HMI tags "DB_SDC_EMS_PAR_DRIVE"
   "_Byte_EMS[XXX].DRIVE_Delay_Pos" : Int, internal   // Absolute Position / absolute Positon
   "_Byte_EMS[XXX].DRIVE_DelaySpeedContr" : Int, internal   // Absolute Position / absolute Positon
   "_Byte_EMS[XXX].DRIVE_DIV_POS_FAST" : Int, internal   // Absolute Position / absolute Positon
   "_Byte_EMS[XXX].DRIVE_DIV_POS_SLOW" : Int, internal   // Absolute Position / absolute Positon
   "_Byte_EMS[XXX].DRIVE_FUNCT" : Int, internal   // Absolute Position / absolute Positon
   "_Byte_EMS[XXX].DRIVE_TOL_RESET_POS" : Int, internal   // Absolute Position / absolute Positon
   "_Byte_EMS[XXX].DRIVE_TOL_SET_POS" : Int, internal   // Absolute Position / absolute Positon
   "_Byte_EMS[XXX].DRIVE_TolSpeedContr" : Int, internal   // Absolute Position / absolute Positon
   "_Byte_EMS[XXX].DRIVE_V_DIV_FAST" : Int, internal   // Absolute Position / absolute Positon
   "_Byte_EMS[XXX].DRIVE_V_FACT_1" : Int, internal   // Absolute Position / absolute Positon
   "_Byte_EMS[XXX].DRIVE_V_FACT_2" : Int, internal   // Absolute Position / absolute Positon
   "_Byte_EMS[XXX].DRIVE_V_FACT_3" : Int, internal   // Absolute Position / absolute Positon
   "_Byte_EMS[XXX].DRIVE_V_FACT_4" : Int, internal   // Absolute Position / absolute Positon
   "_Byte_EMS[XXX].DRIVE_V_FACT_5" : Int, internal   // Absolute Position / absolute Positon
   "_Byte_EMS[XXX].DRIVE_V_Fixed_1" : Int, internal   // Absolute Position / absolute Positon
   "_Byte_EMS[XXX].DRIVE_V_Fixed_2" : Int, internal   // Absolute Position / absolute Positon
   "_Byte_EMS[XXX].DRIVE_V_Fixed_4_SLS_SPEED" : Int, internal   // Absolute Position / absolute Positon
   "_Byte_EMS[XXX].DRIVE_V_LIMIT_FACT" : Int, internal   // Absolute Position / absolute Positon
   "_Byte_EMS[XXX].DRIVE_V_max_Not_top" : Int, internal   // Absolute Position / absolute Positon
   "_Byte_EMS[XXX].DRIVE_V_max_top" : Int, internal   // Absolute Position / absolute Positon
   "_Byte_EMS[XXX].DRIVE_V_min" : Int, internal   // Absolute Position / absolute Positon
   "_Byte_EMS[XXX].DRIVE_V_Pos_2" : Int, internal   // Absolute Position / absolute Positon
   "_Byte_EMS[XXX].DRIVE_V_SETP_1" : Int, internal   // Absolute Position / absolute Positon
   "_Byte_EMS[XXX].DRIVE_V_SETP_2" : Int, internal   // Absolute Position / absolute Positon
   "_Byte_EMS[XXX].DRIVE_V_SETP_3" : Int, internal   // Absolute Position / absolute Positon
   "_Byte_EMS[XXX].DRIVE_V_SETP_4" : Int, internal   // Absolute Position / absolute Positon
   "_Byte_EMS[XXX].DRIVE_Window_Movement" : Int, internal   // Absolute Position / absolute Positon
   "_Byte_EMS[XXX].DRIVE_Window_Overrun" : Int, internal   // Absolute Position / absolute Positon
   "_Byte_EMS[XXX].DRIVE_Window_Pos" : Int, internal   // Absolute Position / absolute Positon
   "_Byte_EMS[XXX].DRIVE_Window_Pos_2" : Int, internal   // Absolute Position / absolute Positon
   "DB_SDC_EMS_PAR_HMI.HMI[XX].PAR.DRIVE.Delay_Pos" : Int AT %DB0.DBW0, 1 s
   "DB_SDC_EMS_PAR_HMI.HMI[XX].PAR.DRIVE.DelaySpeedContr" : S5Time AT %DB0.DBW0, 1 s
   "DB_SDC_EMS_PAR_HMI.HMI[XX].PAR.DRIVE.DIV_POS_FAST" : DInt AT %DB0.DBD0, 1 s
   "DB_SDC_EMS_PAR_HMI.HMI[XX].PAR.DRIVE.DIV_POS_SLOW" : DInt AT %DB0.DBD0, 1 s
   "DB_SDC_EMS_PAR_HMI.HMI[XX].PAR.DRIVE.TOL_RESET_POS" : Int AT %DB0.DBW0, 1 s
   "DB_SDC_EMS_PAR_HMI.HMI[XX].PAR.DRIVE.TOL_SET_POS" : Int AT %DB0.DBW0, 1 s
   "DB_SDC_EMS_PAR_HMI.HMI[XX].PAR.DRIVE.TolSpeedContr" : Int AT %DB0.DBW0, 1 s
   "DB_SDC_EMS_PAR_HMI.HMI[XX].PAR.DRIVE.V_DIV_FAST" : DInt AT %DB0.DBD0, 1 s
   "DB_SDC_EMS_PAR_HMI.HMI[XX].PAR.DRIVE.V_Fixed_1" : DInt AT %DB0.DBD0, 1 s
   "DB_SDC_EMS_PAR_HMI.HMI[XX].PAR.DRIVE.V_Fixed_2" : DInt AT %DB0.DBD0, 1 s
   "DB_SDC_EMS_PAR_HMI.HMI[XX].PAR.DRIVE.V_Fixed_4_SLS_SPEED" : DInt AT %DB0.DBD0, 1 s
   "DB_SDC_EMS_PAR_HMI.HMI[XX].PAR.DRIVE.V_max_Not_top" : DInt AT %DB0.DBD0, 1 s
   "DB_SDC_EMS_PAR_HMI.HMI[XX].PAR.DRIVE.V_max_top" : DInt AT %DB0.DBD0, 1 s
   "DB_SDC_EMS_PAR_HMI.HMI[XX].PAR.DRIVE.V_min" : DInt AT %DB0.DBD0, 1 s
   "DB_SDC_EMS_PAR_HMI.HMI[XX].PAR.DRIVE.V_Pos_2" : DInt AT %DB0.DBD0, 1 s
   "DB_SDC_EMS_PAR_HMI.HMI[XX].PAR.DRIVE.Window_Movement" : Int AT %DB0.DBW0, 1 s
   "DB_SDC_EMS_PAR_HMI.HMI[XX].PAR.DRIVE.Window_Overrun" : Int AT %DB0.DBW0, 1 s
   "DB_SDC_EMS_PAR_HMI.HMI[XX].PAR.DRIVE.Window_Pos" : Int AT %DB0.DBW0, 1 s
   "DB_SDC_EMS_PAR_HMI.HMI[XX].PAR.DRIVE.Window_Pos_2" : Int AT %DB0.DBW0, 1 s
   "DB_SDC_EMS_PAR_HMI.HMI[XX].PAR.DRIVE.Funct" : Word AT %DB0.DBW0, 1 s
   "DB_SDC_EMS_PAR_HMI.HMI[XX].PAR.DRIVE.V_FACT_1" : Real AT %DB0.DBD0, 1 s
   "DB_SDC_EMS_PAR_HMI.HMI[XX].PAR.DRIVE.V_FACT_2" : Real AT %DB0.DBD0, 1 s
   "DB_SDC_EMS_PAR_HMI.HMI[XX].PAR.DRIVE.V_FACT_3" : Real AT %DB0.DBD0, 1 s
   "DB_SDC_EMS_PAR_HMI.HMI[XX].PAR.DRIVE.V_FACT_4" : Real AT %DB0.DBD0, 1 s
   "DB_SDC_EMS_PAR_HMI.HMI[XX].PAR.DRIVE.V_FACT_5" : Real AT %DB0.DBD0, 1 s
   "DB_SDC_EMS_PAR_HMI.HMI[XX].PAR.DRIVE.V_LIMIT_FACT" : Real AT %DB0.DBD0, 1 s
   "DB_SDC_EMS_PAR_HMI.HMI[XX].PAR.DRIVE.V_SETP_1" : DInt AT %DB0.DBD0, 1 s
   "DB_SDC_EMS_PAR_HMI.HMI[XX].PAR.DRIVE.V_SETP_2" : DInt AT %DB0.DBD0, 1 s
   "DB_SDC_EMS_PAR_HMI.HMI[XX].PAR.DRIVE.V_SETP_3" : DInt AT %DB0.DBD0, 1 s
   "DB_SDC_EMS_PAR_HMI.HMI[XX].PAR.DRIVE.V_SETP_4" : DInt AT %DB0.DBD0, 1 s
   "_Byte_EMS[XXX].DRIVE_Delay_Pos(1)" : Int, internal

HMI tags "DB_SDC_EMS_PAR_HOIST"
   "_Byte_EMS[XXX].HOIST_V_min" : Int, internal   // Absolute Position / absolute Positon
   "DB_SDC_EMS_PAR_HMI.HMI[XX].PAR.HOIST.V_min" : Int AT %DB0.DBW0, 1 s
   "_Byte_EMS[XXX].HOIST_V_max" : Int, internal   // Absolute Position / absolute Positon
   "DB_SDC_EMS_PAR_HMI.HMI[XX].PAR.HOIST.V_max" : Int AT %DB0.DBW0, 1 s
   "_Byte_EMS[XXX].HOIST_V_MaxOccLift" : Int, internal   // Absolute Position / absolute Positon
   "DB_SDC_EMS_PAR_HMI.HMI[XX].PAR.HOIST.V_MaxOccLift" : Int AT %DB0.DBW0, 1 s
   "_Byte_EMS[XXX].HOIST_V_Pos_1" : Int, internal   // Absolute Position / absolute Positon
   "DB_SDC_EMS_PAR_HMI.HMI[XX].PAR.HOIST.V_Pos_1" : Int AT %DB0.DBW0, 1 s
   "_Byte_EMS[XXX].HOIST_V_Pos_2" : Int, internal   // Absolute Position / absolute Positon
   "DB_SDC_EMS_PAR_HMI.HMI[XX].PAR.HOIST.V_Pos_2" : Int AT %DB0.DBW0, 1 s
   "_Byte_EMS[XXX].HOIST_V_Fixed_1" : Int, internal   // Absolute Position / absolute Positon
   "DB_SDC_EMS_PAR_HMI.HMI[XX].PAR.HOIST.V_Fixed_1" : Int AT %DB0.DBW0, 1 s
   "_Byte_EMS[XXX].HOIST_V_Fixed_2" : Int, internal   // Absolute Position / absolute Positon
   "DB_SDC_EMS_PAR_HMI.HMI[XX].PAR.HOIST.V_Fixed_2" : Int AT %DB0.DBW0, 1 s
   "_Byte_EMS[XXX].HOIST_V_Fixed_4" : Int, internal   // Absolute Position / absolute Positon
   "DB_SDC_EMS_PAR_HMI.HMI[XX].PAR.HOIST.V_Fixed_4" : Int AT %DB0.DBW0, 1 s
   "_Byte_EMS[XXX].HOIST_V_Fixed_6" : Int, internal   // Absolute Position / absolute Positon
   "DB_SDC_EMS_PAR_HMI.HMI[XX].PAR.HOIST.V_Fixed_6" : Int AT %DB0.DBW0, 1 s
   "_Byte_EMS[XXX].HOIST_V_FACT_Hz_UP" : Int, internal   // Absolute Position / absolute Positon
   "DB_SDC_EMS_PAR_HMI.HMI[XX].PAR.HOIST.V_FACT_Hz_UP" : Real AT %DB0.DBD0, 1 s
   "_Byte_EMS[XXX].HOIST_V_FACT_Hz_DOWN" : Int, internal   // Absolute Position / absolute Positon
   "DB_SDC_EMS_PAR_HMI.HMI[XX].PAR.HOIST.V_FACT_Hz_DOWN" : Real AT %DB0.DBD0, 1 s
   "DB_SDC_EMS_PAR_HMI.HMI[XX].PAR.HOIST.H_Window_POS_V1" : Int AT %DB0.DBW0, 1 s
   "_Byte_EMS[XXX].HOIST_H_Window_POS_V1" : Int, internal   // Absolute Position / absolute Positon
   "DB_SDC_EMS_PAR_HMI.HMI[XX].PAR.HOIST.H_Window_POS_V2" : Int AT %DB0.DBW0, 1 s
   "_Byte_EMS[XXX].HOIST_H_Window_POS_V2" : Int, internal   // Absolute Position / absolute Positon
   "DB_SDC_EMS_PAR_HMI.HMI[XX].PAR.HOIST.H_TOL_SET_POS" : Int AT %DB0.DBW0, 1 s
   "_Byte_EMS[XXX].HOIST_H_TOL_SET_POS" : Int, internal   // Absolute Position / absolute Positon
   "DB_SDC_EMS_PAR_HMI.HMI[XX].PAR.HOIST.H_TOL_RESET_POS" : Int AT %DB0.DBW0, 1 s
   "_Byte_EMS[XXX].HOIST_H_TOL_RESET_POS" : Int, internal   // Absolute Position / absolute Positon
   "DB_SDC_EMS_PAR_HMI.HMI[XX].PAR.HOIST.H_MIN" : Int AT %DB0.DBW0, 1 s
   "_Byte_EMS[XXX].HOIST_H_MIN" : Int, internal   // Absolute Position / absolute Positon
   "DB_SDC_EMS_PAR_HMI.HMI[XX].PAR.HOIST.H_MIN_without_bypass" : Int AT %DB0.DBW0, 1 s
   "_Byte_EMS[XXX].HOIST_H_MIN_without_bypass" : Int, internal   // Absolute Position / absolute Positon
   "DB_SDC_EMS_PAR_HMI.HMI[XX].PAR.HOIST.H_REF_OFFSET" : Int AT %DB0.DBW0, 1 s
   "_Byte_EMS[XXX].HOIST_H_REF_OFFSET" : Int, internal   // Absolute Position / absolute Positon
   "DB_SDC_EMS_PAR_HMI.HMI[XX].PAR.HOIST.H_REF" : Int AT %DB0.DBW0, 1 s
   "_Byte_EMS[XXX].HOIST_H_REF" : Int, internal   // Absolute Position / absolute Positon
   "DB_SDC_EMS_PAR_HMI.HMI[XX].PAR.HOIST.H_FACT_ENC1" : Real AT %DB0.DBD0, 1 s
   "_Byte_EMS[XXX].HOIST_H_FACT_ENC1" : Int, internal   // Absolute Position / absolute Positon
   "DB_SDC_EMS_PAR_HMI.HMI[XX].PAR.HOIST.H_FACT_ENC2" : Real AT %DB0.DBD0, 1 s
   "_Byte_EMS[XXX].HOIST_H_FACT_ENC2" : Int, internal   // Absolute Position / absolute Positon
   "DB_SDC_EMS_PAR_HMI.HMI[XX].PAR.HOIST.H_FACT_SPEED" : Real AT %DB0.DBD0, 1 s
   "_Byte_EMS[XXX].HOIST_H_FACT_SPEED" : Int, internal   // Absolute Position / absolute Positon
   "DB_SDC_EMS_PAR_HMI.HMI[XX].PAR.HOIST.H_ENC_MAX_DIFF" : Int AT %DB0.DBW0, 1 s
   "_Byte_EMS[XXX].HOIST_H_ENC_MAX_DIFF" : Int, internal   // Absolute Position / absolute Positon
   "DB_SDC_EMS_PAR_HMI.HMI[XX].PAR.HOIST.H_Slow" : Int AT %DB0.DBW0, 1 s
   "_Byte_EMS[XXX].HOIST_H_Slow" : Int, internal   // Absolute Position / absolute Positon
   "DB_SDC_EMS_PAR_HMI.HMI[XX].PAR.HOIST.H_tIN_POS" : Int AT %DB0.DBW0, 1 s
   "_Byte_EMS[XXX].HOIST_H_tIN_POS" : Int, internal   // Absolute Position / absolute Positon
   "DB_SDC_EMS_PAR_HMI.HMI[XX].PAR.HOIST.H_REF_HMI" : Int AT %DB0.DBW0, 1 s
   "_Byte_EMS[XXX].HOIST_H_REF_HMI" : Int, internal   // Absolute Position / absolute Positon
   "_Byte_EMS[XXX].HOIST_V_Fixed_3" : Int, internal
   "DB_SDC_EMS_PAR_HMI.HMI[XX].PAR.HOIST.V_Fixed_3" : Int AT %DB0.DBW0, 1 s

HMI tags "VAT_SYSTEM_ALLG"
   "_intern_BILD_Nr" : Int, internal
   "_intern_1_bool" : Bool, internal
   "_intern_0_bool" : Bool, internal
   "_intern_1" : Int, internal
   "_intern_2" : Int, internal
   "_intern_3" : Int, internal
   "_intern_4" : Int, internal
   "_intern_5" : Int, internal
   "_intern_6" : Int, internal
   "_intern_7" : Int, internal
   "_intern_8" : Int, internal
   "_intern_9" : Int, internal
   "_intern_10" : Int, internal
   "_intern_11" : Int, internal
   "_intern_12" : Int, internal
   "_intern_13" : Int, internal
   "_intern_14" : Int, internal
   "_intern_15" : Int, internal
   "_intern_16" : Int, internal
   "_intern_17" : Int, internal
   "_intern_18" : Int, internal
   "_intern_19" : Int, internal
   "_intern_20" : Int, internal
   "_intern_21" : Int, internal
   "_intern_22" : Int, internal
   "_intern_23" : Int, internal
   "_intern_24" : Int, internal
   "_intern_25" : Int, internal
   "_intern_26" : Int, internal
   "_intern_27" : Int, internal
   "_intern_28" : Int, internal
   "_intern_29" : Int, internal
   "_intern_30" : Int, internal
   "_intern_31" : Int, internal
   "_intern_32" : Int, internal
   "_intern_33" : Int, internal
   "_intern_34" : Int, internal
   "_intern_35" : Int, internal
   "_intern_36" : Int, internal
   "_intern_37" : Int, internal
   "_intern_38" : Int, internal
   "_intern_39" : Int, internal
   "_intern_40" : Int, internal
   "_intern_41" : Int, internal
   "_intern_42" : Int, internal
   "_intern_43" : Int, internal
   "_intern_44" : Int, internal
   "_intern_45" : Int, internal
   "_intern_46" : Int, internal
   "_intern_47" : Int, internal
   "_intern_48" : Int, internal
   "_intern_49" : Int, internal
   "_intern_50" : Int, internal
   "_intern_51" : Int, internal
   "_intern_52" : Int, internal
   "_intern_53" : Int, internal
   "_intern_54" : Int, internal
   "_intern_55" : Int, internal
   "_intern_56" : Int, internal
   "_intern_57" : Int, internal
   "_intern_58" : Int, internal
   "_intern_59" : Int, internal
   "_intern_60" : Int, internal
   "_intern_61" : Int, internal
   "_intern_62" : Int, internal
   "_intern_63" : Int, internal
   "_intern_64" : Int, internal
   "_intern_65" : Int, internal
   "_intern_66" : Int, internal
   "_intern_67" : Int, internal
   "_intern_68" : Int, internal
   "_intern_69" : Int, internal
   "_intern_70" : Int, internal
   "_intern_71" : Int, internal
   "_intern_72" : Int, internal
   "_intern_73" : Int, internal
   "_intern_74" : Int, internal
   "_intern_75" : Int, internal
   "_intern_76" : Int, internal
   "_intern_77" : Int, internal
   "_intern_78" : Int, internal
   "_intern_79" : Int, internal
   "_intern_80" : Int, internal
   "_intern_81" : Int, internal
   "_intern_82" : Int, internal
   "_intern_83" : Int, internal
   "_intern_84" : Int, internal
   "_intern_85" : Int, internal
   "_intern_86" : Int, internal
   "_intern_87" : Int, internal
   "_intern_88" : Int, internal
   "_intern_89" : Int, internal
   "_intern_90" : Int, internal
   "_intern_91" : Int, internal
   "_intern_92" : Int, internal
   "_intern_93" : Int, internal
   "_intern_94" : Int, internal
   "_intern_95" : Int, internal
   "_intern_96" : Int, internal
   "_intern_97" : Int, internal
   "_intern_98" : Int, internal
   "_intern_99" : Int, internal
   "_intern_100" : Int, internal
   "_intern_101" : Int, internal
   "_intern_102" : Int, internal
   "_intern_103" : Int, internal
   "_intern_104" : Int, internal
   "_intern_105" : Int, internal
   "_intern_106" : Int, internal
   "_intern_107" : Int, internal
   "_intern_108" : Int, internal
   "_intern_109" : Int, internal
   "_intern_110" : Int, internal
   "_intern_111" : Int, internal
   "_intern_112" : Int, internal
   "_intern_113" : Int, internal
   "_intern_114" : Int, internal
   "_intern_115" : Int, internal
   "_intern_116" : Int, internal
   "_intern_117" : Int, internal
   "_intern_118" : Int, internal
   "_intern_119" : Int, internal
   "_intern_120" : Int, internal
   "_intern_121" : Int, internal
   "_intern_122" : Int, internal
   "_intern_123" : Int, internal
   "_intern_124" : Int, internal
   "_intern_125" : Int, internal
   "_intern_126" : Int, internal
   "_intern_127" : Int, internal
   "_intern_128" : Int, internal
   "_intern_129" : Int, internal
   "_intern_130" : Int, internal
   "_intern_131" : Int, internal
   "_intern_132" : Int, internal
   "_intern_133" : Int, internal
   "_intern_134" : Int, internal
   "_intern_135" : Int, internal
   "_intern_136" : Int, internal
   "_intern_137" : Int, internal
   "_intern_138" : Int, internal
   "_intern_139" : Int, internal
   "_intern_140" : Int, internal
   "_intern_141" : Int, internal
   "_intern_142" : Int, internal
   "_intern_143" : Int, internal
   "_intern_144" : Int, internal
   "_intern_145" : Int, internal
   "_intern_146" : Int, internal
   "_intern_147" : Int, internal
   "_intern_148" : Int, internal
   "_intern_149" : Int, internal
   "_intern_150" : Int, internal
   "_intern_151" : Int, internal
   "_intern_152" : Int, internal
   "_intern_153" : Int, internal
   "_intern_154" : Int, internal
   "_intern_155" : Int, internal
   "_intern_156" : Int, internal
   "_intern_157" : Int, internal
   "_intern_158" : Int, internal
   "_intern_159" : Int, internal
   "_intern_160" : Int, internal
   "_intern_161" : Int, internal
   "_intern_162" : Int, internal
   "_intern_163" : Int, internal
   "_intern_164" : Int, internal
   "_intern_165" : Int, internal
   "_intern_166" : Int, internal
   "_intern_167" : Int, internal
   "_intern_168" : Int, internal
   "_intern_169" : Int, internal
   "_intern_170" : Int, internal
   "_intern_171" : Int, internal
   "_intern_172" : Int, internal
   "_intern_173" : Int, internal
   "_intern_174" : Int, internal
   "_intern_175" : Int, internal
   "_intern_176" : Int, internal
   "_intern_177" : Int, internal
   "_intern_178" : Int, internal
   "_intern_179" : Int, internal
   "_intern_180" : Int, internal
   "_intern_181" : Int, internal
   "_intern_182" : Int, internal
   "_intern_183" : Int, internal
   "_intern_184" : Int, internal
   "_intern_185" : Int, internal
   "_intern_186" : Int, internal
   "_intern_187" : Int, internal
   "_intern_188" : Int, internal
   "_intern_189" : Int, internal
   "_intern_190" : Int, internal
   "_intern_191" : Int, internal
   "_intern_192" : Int, internal
   "_intern_193" : Int, internal
   "_intern_194" : Int, internal
   "_intern_195" : Int, internal
   "_intern_196" : Int, internal
   "_intern_197" : Int, internal
   "_intern_198" : Int, internal
   "_intern_199" : Int, internal
   "_intern_200" : Int, internal

HMI tags "VAT_PN_PB"
   "PN_PB\PTMUX_P_TLN17_32" : UInt, internal
   "PN_PB\PTMUX_P_TLN1_16" : UInt, internal
   "PN_PB\PTMUX_P_TLN129_144" : UInt, internal
   "PN_PB\DB_PN" : UInt, internal
   "PN_PB\PTMUX_P_TLN177_192" : UInt, internal
   "PN_PB\PTMUX_F_TLN241_256" : UInt, internal
   "PN_PB\IO_Sys_ID" : Int, internal
   "PN_PB\PTMUX_P_TLN225_240" : UInt, internal
   "PN_PB\PTMUX_P_TLN241_256" : UInt, internal
   "PN_PB\PTMUX_P_TLN193_208" : UInt, internal
   "PN_PB\PTMUX_F_TLN1_16" : UInt, internal
   "PN_PB\PTMUX_P_TLN209_224" : UInt, internal
   "PN_PB\PTMUX_F_TLN49_64" : UInt, internal
   "PN_PB\PTMUX_P_TLN113_128" : UInt, internal
   "PN_PB\PTMUX_F_TLN177_192" : UInt, internal
   "PN_PB\PTMUX_P_TLN49_64" : UInt, internal
   "PN_PB\PTMUX_F_TLN97_112" : UInt, internal
   "PN_PB\DB_PB" : UInt, internal
   "PN_PB\PTMUX_F_TLN81_96" : UInt, internal
   "PN_PB\PTMUX_F_TLN145_160" : UInt, internal
   "PN_PB\Diag_Art" : Int, internal
   "PN_PB\PTMUX_F_TLN113_128" : UInt, internal
   "PN_PB\PTMUX_P_TLN97_112" : UInt, internal
   "PN_PB\Teiln_Nr_Anz." : Int, internal
   "PN_PB\PTMUX_P_TLN33_48" : UInt, internal
   "PN_PB\PTMUX_F_TLN161_176" : UInt, internal
   "PN_PB\PTMUX_F_TLN193_208" : UInt, internal
   "PN_PB\PTMUX_P_TLN81_96" : UInt, internal
   "PN_PB\PTMUX_P_TLN65_80" : UInt, internal
   "PN_PB\PTMUX_F_TLN225_240" : UInt, internal
   "PN_PB\PTMUX_F_TLN17_32" : UInt, internal
   "PN_PB\PTMUX_F_TLN65_80" : UInt, internal
   "PN_PB\PTMUX_F_TLN209_224" : UInt, internal
   "PN_PB\PTMUX_F_TLN33_48" : UInt, internal
   "PN_PB\PTMUX_P_TLN145_160" : UInt, internal
   "PN_PB\PTMUX_P_TLN161_176" : UInt, internal
   "PN_PB\Teiln_Nr_Bez" : WString[20], internal
   "PN_PB\Teiln_Nr_Typ" : WString[12], internal
   "PN_PB\Teiln_Nr_Ort" : WString[12], internal
   "PN_PB\PTMUX_F_TLN129_144" : UInt, internal

HMI tags "VAT_SYSTEM_PN"
   "PN_PB\PN\TLN_P_161_176" : Word AT %DB0.DBW230, 100 ms
   "PN_PB\PN\TLN_F_241_256" : Word AT %DB0.DBW368, 100 ms
   "PN_PB\PN\TLN_P_33_48" : Word AT %DB0.DBW214, 100 ms
   "PN_PB\PN\TLN_F_49_64" : Word AT %DB0.DBW344, 100 ms
   "PN_PB\PN\TLN_F_81_96" : Word AT %DB0.DBW348, 100 ms
   "PN_PB\PN\TLN_P_225_240" : Word AT %DB0.DBW238, 100 ms
   "PN_PB\PN\TLN_P_177_192" : Word AT %DB0.DBW232, 100 ms
   "PN_PB\PN\TLN_F_17_32" : Word AT %DB0.DBW340, 100 ms
   "PN_PB\PN\TLN_F_225_240" : Word AT %DB0.DBW366, 100 ms
   "PN_PB\PN\TLN_F_33_48" : Word AT %DB0.DBW342, 100 ms
   "PN_PB\PN\TLN_P_97_112" : Word AT %DB0.DBW222, 100 ms
   "PN_PB\PN\TLN_P_129_144" : Word AT %DB0.DBW226, 100 ms
   "PN_PB\PN\Diag_Slave_Nr" : Int, internal
   "PN_PB\PN\TLN_F_113_128" : Word AT %DB0.DBW352, 100 ms
   "PN_PB\PN\TLN_F_97_112" : Word AT %DB0.DBW350, 100 ms
   "PN_PB\PN\TLN_P_145_160" : Word AT %DB0.DBW228, 100 ms
   "PN_PB\PN\TLN_F_145_160" : Word AT %DB0.DBW356, 100 ms
   "PN_PB\PN\TLN_P_113_128" : Word AT %DB0.DBW224, 100 ms
   "PN_PB\PN\IOSys_ID" : Int AT %DB0.DBW2, 200 ms
   "PN_PB\PN\TLN_F_129_144" : Word AT %DB0.DBW354, 100 ms
   "PN_PB\PN\TLN_F_161_176" : Word AT %DB0.DBW358, 100 ms
   "PN_PB\PN\TLN_F_1_16" : Word AT %DB0.DBW338, 100 ms
   "PN_PB\PN\TLN_P_1_16" : Word AT %DB0.DBW210, 100 ms
   "PN_PB\PN\TLN_P_65_80" : Word AT %DB0.DBW218, 100 ms
   "PN_PB\PN\TLN_F_209_224" : Word AT %DB0.DBW364, 100 ms
   "PN_PB\PN\TLN_F_65_80" : Word AT %DB0.DBW346, 100 ms
   "PN_PB\PN\TLN_P_193_208" : Word AT %DB0.DBW234, 100 ms
   "PN_PB\PN\TLN_P_81_96" : Word AT %DB0.DBW220, 100 ms
   "PN_PB\PN\TLN_P_209_224" : Word AT %DB0.DBW236, 100 ms
   "PN_PB\PN\TLN_P_17_32" : Word AT %DB0.DBW212, 100 ms
   "PN_PB\PN\TLN_P_49_64" : Word AT %DB0.DBW216, 100 ms
   "PN_PB\PN\TLN_P_241_256" : Word AT %DB0.DBW240, 100 ms
   "PN_PB\PN\TLN_F_193_208" : Word AT %DB0.DBW362, 100 ms
   "PN_PB\PN\TLN_F_177_192" : Word AT %DB0.DBW360, 100 ms
   "PN_PB\PN\Teiln_Nr" : Int AT %DB0.DBW4, 1 s
      on ChangeValue: "SDC_PN"()

HMI tags "VAT_SYSTEM_PB"
   "PN_PB\PB\TLN_F_65_80" : Word AT %DB0.DBW234, 100 ms
   "PN_PB\PB\TLN_F_113_128" : Word AT %DB0.DBW240, 100 ms
   "PN_PB\PB\IOSys_ID" : Int AT %DB0.DBW2, 200 ms
   "PN_PB\PB\TLN_P_81_96" : Word AT %DB0.DBW220, 100 ms
   "PN_PB\PB\TLN_F_81_96" : Word AT %DB0.DBW236, 100 ms
   "PN_PB\PB\TLN_F_49_64" : Word AT %DB0.DBW232, 100 ms
   "PN_PB\PB\TLN_P_113_128" : Word AT %DB0.DBW224, 100 ms
   "PN_PB\PB\TLN_F_33_48" : Word AT %DB0.DBW230, 100 ms
   "PN_PB\PB\TLN_P_65_80" : Word AT %DB0.DBW218, 100 ms
   "PN_PB\PB\TLN_P_49_64" : Word AT %DB0.DBW216, 100 ms
   "PN_PB\PB\TLN_F_1_16" : Word AT %DB0.DBW226, 100 ms
   "PN_PB\PB\TLN_P_17_32" : Word AT %DB0.DBW212, 100 ms
   "PN_PB\PB\TLN_P_33_48" : Word AT %DB0.DBW214, 100 ms
   "PN_PB\PB\TLN_P_1_16" : Word AT %DB0.DBW210, 100 ms
   "PN_PB\PB\TLN_F_17_32" : Word AT %DB0.DBW228, 100 ms
   "PN_PB\PB\TLN_F_97_112" : Word AT %DB0.DBW238, 100 ms
   "PN_PB\PB\TLN_P_97_112" : Word AT %DB0.DBW222, 100 ms
   "PN_PB\PB\Teiln_Nr" : Int AT %DB0.DBW4, 200 ms

HMI tags "VAT_SYSTEM_PARAMETER"
   "_intern_Pult_Nr" : Int, internal   // !!! VOR DEM LADEN EINSTELLEN !!!

HMI tags "UserDiag_TagTable"
   "UserDiag_HmiData_actIOSystem" : Int = PLC UserDiag_HmiData.actIOSystem, 1 s
   "UserDiag_HmiData_actDeviceOfScreen" : Int = PLC UserDiag_HmiData.actDeviceOfScreen, 1 s
   "UserDiag_HmiData_ioSlotDiagnosticsLoaded" : Bool = PLC UserDiag_HmiData.ioSlotDiagnosticsLoaded, 1 s
   "UserDiag_HmiData_actScreenDevices" : Int = PLC UserDiag_HmiData.actScreenDevices, 100 ms
   "UserDiag_HmiData_maxScreensDevices" : Int = PLC UserDiag_HmiData.maxScreensDevices, 1 s
   "UserDiag_HmiData_ackWaitTime" : Int = PLC UserDiag_HmiData.ackWaitTime, 1 s
   "UserDiag_HmiData_ackStates" : Bool = PLC UserDiag_HmiData.ackStates, 1 s
   "UserDiag_HmiData_actIOSystemData" : UserDiag_typeActIOSystem = PLC UserDiag_HmiData.actIOSystemData, 1 s
   "UserDiag_HmiData_actDeviceNumber" : UInt = PLC UserDiag_HmiData.actDeviceNumber, 1 s
   "UserDiag_HmiData_actDeviceName" : String[50] = PLC UserDiag_HmiData.actDeviceName, 1 s
   "UserDiag_HmiData_actIPAddress.ADDR" : Array [0..3] of Byte = PLC UserDiag_HmiData.actIPAddress.ADDR, 1 s
   "UserDiag_HmiData_ioSystemError" : Array [0..1] of Bool = PLC UserDiag_HmiData.ioSystemError AT %DB1.DBX0.0, 500 ms
   "UserDiag_HmiData_filterErrorDevices" : Bool = PLC UserDiag_HmiData.filterErrorDevices AT %DB1.DBX0.0, 500 ms
   "UserDiag_HmiData_errorAtLowerScreen" : Bool = PLC UserDiag_HmiData.errorAtLowerScreen, 500 ms
   "UserDiag_HmiData_errorAtUpperScreen" : Bool = PLC UserDiag_HmiData.errorAtUpperScreen AT %DB1.DBW0, 500 ms
   "ioSystem1" : Int AT %DB1.DBW0
   "ioSystem2" : Int AT %DB1.DBW0
   "ioSystem3" : Int AT %DB1.DBW0
   "DB_SDC_FAULTS" : Word = PLC DB101_DB_SDC_FAULTS.SDC_Fault AT %DB101.DBW0, 1 s

HMI tags "DB_SDC_FAULTS"
   "DB101_DB_SDC_FAULTS_SDC_Fault" : Word = PLC DB101_DB_SDC_FAULTS.SDC_Fault AT %DB101.DBW0, 1 s
   "DB101_DB_SDC_FAULTS_Carrier_Fault[15]" : Word = PLC DB101_DB_SDC_FAULTS.Carrier_Fault[15] AT %DB101.DBW30, 1 s
   "DB101_DB_SDC_FAULTS_Carrier_Fault[27]" : Word = PLC DB101_DB_SDC_FAULTS.Carrier_Fault[27] AT %DB101.DBW54, 1 s
   "DB101_DB_SDC_FAULTS_Carrier_Fault[31]" : Word = PLC DB101_DB_SDC_FAULTS.Carrier_Fault[31] AT %DB101.DBW62, 1 s
   "DB101_DB_SDC_FAULTS_Carrier_Fault[40]" : Word = PLC DB101_DB_SDC_FAULTS.Carrier_Fault[40] AT %DB101.DBW80, 1 s

HMI tags "DB_HMI_FAULTS"
   "DB302_HMI_Faults_SDC_Faults_0" : Int = PLC DB302_HMI_Faults.SDC_Faults_0, 1 s
   "DB302_HMI_Faults_SDC_Faults_1" : Int = PLC DB302_HMI_Faults.SDC_Faults_1, 1 s
   "DB302_HMI_Faults_SDC_Faults_2" : Int = PLC DB302_HMI_Faults.SDC_Faults_2, 1 s
   "DB302_HMI_Faults_SDC_Faults_3" : Int = PLC DB302_HMI_Faults.SDC_Faults_3, 1 s

HMI tags "EMS"
   "EMS" : UDT_System = PLC EMS AT %DB1.DBW0, 1 s

HMI tags "DeviceStates_Condition"
   "DB16_EMS_Status_EMS_DeviceStates.DeviceStates_Condition_HMI[2]" : Int = PLC DB16_EMS_Status.EMS_DeviceStates.DeviceStates_Condition_HMI[2], 1 s
   "DB16_EMS_Status_EMS_DeviceStates.DeviceStates_Condition_HMI[3]" : Int = PLC DB16_EMS_Status.EMS_DeviceStates.DeviceStates_Condition_HMI[3], 1 s
   "DB16_EMS_Status_EMS_DeviceStates.DeviceStates_Condition_HMI[4]" : Int = PLC DB16_EMS_Status.EMS_DeviceStates.DeviceStates_Condition_HMI[4], 1 s
   "DB16_EMS_Status_EMS_DeviceStates.DeviceStates_Condition_HMI[5]" : Int = PLC DB16_EMS_Status.EMS_DeviceStates.DeviceStates_Condition_HMI[5], 1 s
   "DB16_EMS_Status_EMS_DeviceStates.DeviceStates_Condition_HMI[6]" : Int = PLC DB16_EMS_Status.EMS_DeviceStates.DeviceStates_Condition_HMI[6], 1 s
   "DB16_EMS_Status_EMS_DeviceStates.DeviceStates_Condition_HMI[7]" : Int = PLC DB16_EMS_Status.EMS_DeviceStates.DeviceStates_Condition_HMI[7], 1 s
   "DB16_EMS_Status_EMS_DeviceStates.DeviceStates_Condition_HMI[8]" : Int = PLC DB16_EMS_Status.EMS_DeviceStates.DeviceStates_Condition_HMI[8], 1 s
   "DB16_EMS_Status_EMS_DeviceStates.DeviceStates_Condition_HMI[9]" : Int = PLC DB16_EMS_Status.EMS_DeviceStates.DeviceStates_Condition_HMI[9], 1 s
   "DB16_EMS_Status_EMS_DeviceStates.DeviceStates_Condition_HMI[10]" : Int = PLC DB16_EMS_Status.EMS_DeviceStates.DeviceStates_Condition_HMI[10], 1 s
   "DB16_EMS_Status_EMS_DeviceStates.DeviceStates_Condition_HMI[11]" : Int = PLC DB16_EMS_Status.EMS_DeviceStates.DeviceStates_Condition_HMI[11], 1 s
   "DB16_EMS_Status_EMS_DeviceStates.DeviceStates_Condition_HMI[12]" : Int = PLC DB16_EMS_Status.EMS_DeviceStates.DeviceStates_Condition_HMI[12], 1 s
   "DB16_EMS_Status_EMS_DeviceStates.DeviceStates_Condition_HMI[13]" : Int = PLC DB16_EMS_Status.EMS_DeviceStates.DeviceStates_Condition_HMI[13], 1 s
   "DB16_EMS_Status_EMS_DeviceStates.DeviceStates_Condition_HMI[14]" : Int = PLC DB16_EMS_Status.EMS_DeviceStates.DeviceStates_Condition_HMI[14], 1 s
   "DB16_EMS_Status_EMS_DeviceStates.DeviceStates_Condition_HMI[15]" : Int = PLC DB16_EMS_Status.EMS_DeviceStates.DeviceStates_Condition_HMI[15], 1 s
   "DB16_EMS_Status_EMS_DeviceStates.DeviceStates_Condition_HMI[16]" : Int = PLC DB16_EMS_Status.EMS_DeviceStates.DeviceStates_Condition_HMI[16], 1 s
   "DB16_EMS_Status_EMS_DeviceStates.DeviceStates_Condition_HMI[17]" : Int = PLC DB16_EMS_Status.EMS_DeviceStates.DeviceStates_Condition_HMI[17], 1 s
   "DB16_EMS_Status_EMS_DeviceStates.DeviceStates_Condition_HMI[18]" : Int = PLC DB16_EMS_Status.EMS_DeviceStates.DeviceStates_Condition_HMI[18], 1 s
   "DB16_EMS_Status_EMS_DeviceStates.DeviceStates_Condition_HMI[19]" : Int = PLC DB16_EMS_Status.EMS_DeviceStates.DeviceStates_Condition_HMI[19], 1 s
   "DB16_EMS_Status_EMS_DeviceStates.DeviceStates_Condition_HMI[20]" : Int = PLC DB16_EMS_Status.EMS_DeviceStates.DeviceStates_Condition_HMI[20], 1 s
   "DB16_EMS_Status_EMS_DeviceStates.DeviceStates_Condition_HMI[21]" : Int = PLC DB16_EMS_Status.EMS_DeviceStates.DeviceStates_Condition_HMI[21], 1 s
   "DB16_EMS_Status_EMS_DeviceStates.DeviceStates_Condition_HMI[22]" : Int = PLC DB16_EMS_Status.EMS_DeviceStates.DeviceStates_Condition_HMI[22], 1 s
   "DB16_EMS_Status_EMS_DeviceStates.DeviceStates_Condition_HMI[23]" : Int = PLC DB16_EMS_Status.EMS_DeviceStates.DeviceStates_Condition_HMI[23], 1 s
   "DB16_EMS_Status_EMS_DeviceStates.DeviceStates_Condition_HMI[24]" : Int = PLC DB16_EMS_Status.EMS_DeviceStates.DeviceStates_Condition_HMI[24], 1 s
   "DB16_EMS_Status_EMS_DeviceStates.DeviceStates_Condition_HMI[25]" : Int = PLC DB16_EMS_Status.EMS_DeviceStates.DeviceStates_Condition_HMI[25], 1 s
   "DB16_EMS_Status_EMS_DeviceStates.DeviceStates_Condition_HMI[26]" : Int = PLC DB16_EMS_Status.EMS_DeviceStates.DeviceStates_Condition_HMI[26], 1 s
   "DB16_EMS_Status_EMS_DeviceStates.DeviceStates_Condition_HMI[27]" : Int = PLC DB16_EMS_Status.EMS_DeviceStates.DeviceStates_Condition_HMI[27], 1 s
   "DB16_EMS_Status_EMS_DeviceStates.DeviceStates_Condition_HMI[28]" : Int = PLC DB16_EMS_Status.EMS_DeviceStates.DeviceStates_Condition_HMI[28], 1 s
   "DB16_EMS_Status_EMS_DeviceStates.DeviceStates_Condition_HMI[29]" : Int = PLC DB16_EMS_Status.EMS_DeviceStates.DeviceStates_Condition_HMI[29], 1 s
   "DB16_EMS_Status_EMS_DeviceStates.DeviceStates_Condition_HMI[30]" : Int = PLC DB16_EMS_Status.EMS_DeviceStates.DeviceStates_Condition_HMI[30], 1 s
   "DB16_EMS_Status_EMS_DeviceStates.DeviceStates_Condition_HMI[31]" : Int = PLC DB16_EMS_Status.EMS_DeviceStates.DeviceStates_Condition_HMI[31], 1 s
   "DB16_EMS_Status_EMS_DeviceStates.DeviceStates_Condition_HMI[32]" : Int = PLC DB16_EMS_Status.EMS_DeviceStates.DeviceStates_Condition_HMI[32], 1 s
   "DB16_EMS_Status_EMS_DeviceStates.DeviceStates_Condition_HMI[33]" : Int = PLC DB16_EMS_Status.EMS_DeviceStates.DeviceStates_Condition_HMI[33], 1 s
   "DB16_EMS_Status_EMS_DeviceStates.DeviceStates_Condition_HMI[34]" : Int = PLC DB16_EMS_Status.EMS_DeviceStates.DeviceStates_Condition_HMI[34], 1 s
   "DB16_EMS_Status_EMS_DeviceStates.DeviceStates_Condition_HMI[35]" : Int = PLC DB16_EMS_Status.EMS_DeviceStates.DeviceStates_Condition_HMI[35], 1 s
   "DB16_EMS_Status_EMS_DeviceStates.DeviceStates_Condition_HMI[36]" : Int = PLC DB16_EMS_Status.EMS_DeviceStates.DeviceStates_Condition_HMI[36], 1 s
   "DB16_EMS_Status_EMS_DeviceStates.DeviceStates_Condition_HMI[37]" : Int = PLC DB16_EMS_Status.EMS_DeviceStates.DeviceStates_Condition_HMI[37], 1 s
   "DB16_EMS_Status_EMS_DeviceStates.DeviceStates_Condition_HMI[38]" : Int = PLC DB16_EMS_Status.EMS_DeviceStates.DeviceStates_Condition_HMI[38], 1 s
   "DB16_EMS_Status_EMS_DeviceStates.DeviceStates_Condition_HMI[39]" : Int = PLC DB16_EMS_Status.EMS_DeviceStates.DeviceStates_Condition_HMI[39], 1 s
   "DB16_EMS_Status_EMS_DeviceStates.DeviceStates_Condition_HMI[40]" : Int = PLC DB16_EMS_Status.EMS_DeviceStates.DeviceStates_Condition_HMI[40], 1 s
   "DB16_EMS_Status_EMS_DeviceStates.DeviceStates_Condition_HMI[41]" : Int = PLC DB16_EMS_Status.EMS_DeviceStates.DeviceStates_Condition_HMI[41], 1 s
   "DB16_EMS_Status_EMS_DeviceStates.DeviceStates_Condition_HMI[42]" : Int = PLC DB16_EMS_Status.EMS_DeviceStates.DeviceStates_Condition_HMI[42], 1 s
   "DB16_EMS_Status_EMS_DeviceStates.DeviceStates_Condition_HMI[43]" : Int = PLC DB16_EMS_Status.EMS_DeviceStates.DeviceStates_Condition_HMI[43], 1 s
   "DB16_EMS_Status_EMS_DeviceStates.DeviceStates_Condition_HMI[44]" : Int = PLC DB16_EMS_Status.EMS_DeviceStates.DeviceStates_Condition_HMI[44], 1 s
   "DB16_EMS_Status_EMS_DeviceStates.DeviceStates_Condition_HMI[45]" : Int = PLC DB16_EMS_Status.EMS_DeviceStates.DeviceStates_Condition_HMI[45], 1 s
   "DB16_EMS_Status_EMS_DeviceStates.DeviceStates_Condition_HMI[46]" : Int = PLC DB16_EMS_Status.EMS_DeviceStates.DeviceStates_Condition_HMI[46], 1 s
   "DB16_EMS_Status_EMS_DeviceStates.DeviceStates_Condition_HMI[47]" : Int = PLC DB16_EMS_Status.EMS_DeviceStates.DeviceStates_Condition_HMI[47], 1 s
   "DB16_EMS_Status_EMS_DeviceStates.DeviceStates_Condition_HMI[48]" : Int = PLC DB16_EMS_Status.EMS_DeviceStates.DeviceStates_Condition_HMI[48], 1 s
   "DB16_EMS_Status_EMS_DeviceStates.DeviceStates_Condition_HMI[49]" : Int = PLC DB16_EMS_Status.EMS_DeviceStates.DeviceStates_Condition_HMI[49], 1 s
   "DB16_EMS_Status_EMS_DeviceStates.DeviceStates_Condition_HMI[50]" : Int = PLC DB16_EMS_Status.EMS_DeviceStates.DeviceStates_Condition_HMI[50], 1 s
   "DB16_EMS_Status_EMS_DeviceStates.DeviceStates_Condition_HMI[51]" : Int = PLC DB16_EMS_Status.EMS_DeviceStates.DeviceStates_Condition_HMI[51], 1 s
   "DB16_EMS_Status_EMS_DeviceStates.DeviceStates_Condition_HMI[52]" : Int = PLC DB16_EMS_Status.EMS_DeviceStates.DeviceStates_Condition_HMI[52], 1 s
   "DB16_EMS_Status_EMS_DeviceStates.DeviceStates_Condition_HMI[53]" : Int = PLC DB16_EMS_Status.EMS_DeviceStates.DeviceStates_Condition_HMI[53], 1 s
   "DB16_EMS_Status_EMS_DeviceStates.DeviceStates_Condition_HMI[54]" : Int = PLC DB16_EMS_Status.EMS_DeviceStates.DeviceStates_Condition_HMI[54], 1 s
   "DB16_EMS_Status_EMS_DeviceStates.DeviceStates_Condition_HMI[55]" : Int = PLC DB16_EMS_Status.EMS_DeviceStates.DeviceStates_Condition_HMI[55], 1 s
   "DB16_EMS_Status_EMS_DeviceStates.DeviceStates_Condition_HMI[56]" : Int = PLC DB16_EMS_Status.EMS_DeviceStates.DeviceStates_Condition_HMI[56], 1 s
   "DB16_EMS_Status_EMS_DeviceStates.DeviceStates_Condition_HMI[57]" : Int = PLC DB16_EMS_Status.EMS_DeviceStates.DeviceStates_Condition_HMI[57], 1 s
   "DB16_EMS_Status_EMS_DeviceStates.DeviceStates_Condition_HMI[58]" : Int = PLC DB16_EMS_Status.EMS_DeviceStates.DeviceStates_Condition_HMI[58], 1 s
   "DB16_EMS_Status_EMS_DeviceStates.DeviceStates_Condition_HMI[59]" : Int = PLC DB16_EMS_Status.EMS_DeviceStates.DeviceStates_Condition_HMI[59], 1 s
   "DB16_EMS_Status_EMS_DeviceStates.DeviceStates_Condition_HMI[60]" : Int = PLC DB16_EMS_Status.EMS_DeviceStates.DeviceStates_Condition_HMI[60], 1 s
   "DB16_EMS_Status_EMS_DeviceStates.DeviceStates_Condition_HMI[61]" : Int = PLC DB16_EMS_Status.EMS_DeviceStates.DeviceStates_Condition_HMI[61], 1 s
   "DB16_EMS_Status_EMS_DeviceStates.DeviceStates_Condition_HMI[62]" : Int = PLC DB16_EMS_Status.EMS_DeviceStates.DeviceStates_Condition_HMI[62], 1 s
   "DB16_EMS_Status_EMS_DeviceStates.DeviceStates_Condition_HMI[63]" : Int = PLC DB16_EMS_Status.EMS_DeviceStates.DeviceStates_Condition_HMI[63], 1 s
   "DB16_EMS_Status_EMS_DeviceStates.DeviceStates_Condition_HMI[64]" : Int = PLC DB16_EMS_Status.EMS_DeviceStates.DeviceStates_Condition_HMI[64], 1 s
   "DB16_EMS_Status_EMS_DeviceStates.DeviceStates_Condition_HMI[65]" : Int = PLC DB16_EMS_Status.EMS_DeviceStates.DeviceStates_Condition_HMI[65], 1 s
   "DB16_EMS_Status_EMS_DeviceStates.DeviceStates_Condition_HMI[66]" : Int = PLC DB16_EMS_Status.EMS_DeviceStates.DeviceStates_Condition_HMI[66], 1 s
   "DB16_EMS_Status_EMS_DeviceStates.DeviceStates_Condition_HMI[67]" : Int = PLC DB16_EMS_Status.EMS_DeviceStates.DeviceStates_Condition_HMI[67], 1 s
   "DB16_EMS_Status_EMS_DeviceStates.DeviceStates_Condition_HMI[68]" : Int = PLC DB16_EMS_Status.EMS_DeviceStates.DeviceStates_Condition_HMI[68], 1 s
   "DB16_EMS_Status_EMS_DeviceStates.DeviceStates_Condition_HMI[69]" : Int = PLC DB16_EMS_Status.EMS_DeviceStates.DeviceStates_Condition_HMI[69], 1 s
   "DB16_EMS_Status_EMS_DeviceStates.DeviceStates_Condition_HMI[70]" : Int = PLC DB16_EMS_Status.EMS_DeviceStates.DeviceStates_Condition_HMI[70], 1 s
   "DB16_EMS_Status_EMS_DeviceStates.DeviceStates_Condition_HMI[71]" : Int = PLC DB16_EMS_Status.EMS_DeviceStates.DeviceStates_Condition_HMI[71], 1 s
   "DB16_EMS_Status_EMS_DeviceStates.DeviceStates_Condition_HMI[72]" : Int = PLC DB16_EMS_Status.EMS_DeviceStates.DeviceStates_Condition_HMI[72], 1 s
   "DB16_EMS_Status_EMS_DeviceStates.DeviceStates_Condition_HMI[73]" : Int = PLC DB16_EMS_Status.EMS_DeviceStates.DeviceStates_Condition_HMI[73], 1 s
   "DB16_EMS_Status_EMS_DeviceStates.DeviceStates_Condition_HMI[74]" : Int = PLC DB16_EMS_Status.EMS_DeviceStates.DeviceStates_Condition_HMI[74], 1 s
   "DB16_EMS_Status_EMS_DeviceStates.DeviceStates_Condition_HMI[75]" : Int = PLC DB16_EMS_Status.EMS_DeviceStates.DeviceStates_Condition_HMI[75], 1 s
   "DB16_EMS_Status_EMS_DeviceStates.DeviceStates_Condition_HMI[76]" : Int = PLC DB16_EMS_Status.EMS_DeviceStates.DeviceStates_Condition_HMI[76], 1 s
   "DB16_EMS_Status_EMS_DeviceStates.DeviceStates_Condition_HMI[77]" : Int = PLC DB16_EMS_Status.EMS_DeviceStates.DeviceStates_Condition_HMI[77], 1 s
   "DB16_EMS_Status_EMS_DeviceStates.DeviceStates_Condition_HMI[78]" : Int = PLC DB16_EMS_Status.EMS_DeviceStates.DeviceStates_Condition_HMI[78], 1 s
   "DB16_EMS_Status_EMS_DeviceStates.DeviceStates_Condition_HMI[79]" : Int = PLC DB16_EMS_Status.EMS_DeviceStates.DeviceStates_Condition_HMI[79], 1 s
   "DB16_EMS_Status_EMS_DeviceStates.DeviceStates_Condition_HMI[80]" : Int = PLC DB16_EMS_Status.EMS_DeviceStates.DeviceStates_Condition_HMI[80], 1 s
   "DB16_EMS_Status_EMS_DeviceStates.DeviceStates_Condition_HMI[81]" : Int = PLC DB16_EMS_Status.EMS_DeviceStates.DeviceStates_Condition_HMI[81], 1 s
   "DB16_EMS_Status_EMS_DeviceStates.DeviceStates_Condition_HMI[82]" : Int = PLC DB16_EMS_Status.EMS_DeviceStates.DeviceStates_Condition_HMI[82], 1 s
   "DB16_EMS_Status_EMS_DeviceStates.DeviceStates_Condition_HMI[1]" : Int = PLC DB16_EMS_Status.EMS_DeviceStates.DeviceStates_Condition_HMI[1], 1 s
   "DB16_EMS_Status_EMS_DeviceStates.DeviceStates_Condition_HMI" : Array [0..82] of Int = PLC DB16_EMS_Status.EMS_DeviceStates.DeviceStates_Condition_HMI AT %DB1.DBW0, 1 s

